   		
   		'KANAN
   		b21d3eaf-4e31-425c-ad1a-ba4e4002cacc Tool_Allocation_Numb_16,76
   		b21d3eaf-4e31-425c-ad1a-ba4e4002cacc Tool_Allocation_Numb_17,77
   		b21d3eaf-4e31-425c-ad1a-ba4e4002cacc Tool_Allocation_Numb_18,78
   		b21d3eaf-4e31-425c-ad1a-ba4e4002cacc Tool_Allocation_Numb_19,79
   		b21d3eaf-4e31-425c-ad1a-ba4e4002cacc Tool_Allocation_Numb_20,80
   		b21d3eaf-4e31-425c-ad1a-ba4e4002cacc Tool_Allocation_Numb_21,81
   		b21d3eaf-4e31-425c-ad1a-ba4e4002cacc Tool_Allocation_Numb_22,82
   		b21d3eaf-4e31-425c-ad1a-ba4e4002cacc Tool_Allocation_Numb_23,83
   		b21d3eaf-4e31-425c-ad1a-ba4e4002cacc Tool_Allocation_Numb_24,84
   		b21d3eaf-4e31-425c-ad1a-ba4e4002cacc Tool_Allocation_Numb_25,85
   		b21d3eaf-4e31-425c-ad1a-ba4e4002cacc Tool_Allocation_Numb_26,86
   		b21d3eaf-4e31-425c-ad1a-ba4e4002cacc Tool_Allocation_Numb_27,87
   		b21d3eaf-4e31-425c-ad1a-ba4e4002cacc Tool_Allocation_Numb_28,88
   		b21d3eaf-4e31-425c-ad1a-ba4e4002cacc Tool_Allocation_Numb_29,89
   		b21d3eaf-4e31-425c-ad1a-ba4e4002cacc Tool_Allocation_Numb_30,90		
   Case 4
   		b21d3eaf-4e31-425c-ad1a-ba4e4002cacc Tool_Allocation_Numb_1,91
   		b21d3eaf-4e31-425c-ad1a-ba4e4002cacc Tool_Allocation_Numb_2,92
   		b21d3eaf-4e31-425c-ad1a-ba4e4002cacc Tool_Allocation_Numb_3,93
   		b21d3eaf-4e31-425c-ad1a-ba4e4002cacc Tool_Allocation_Numb_4,94
   		b21d3eaf-4e31-425c-ad1a-ba4e4002cacc Tool_Allocation_Numb_5,95
   		b21d3eaf-4e31-425c-ad1a-ba4e4002cacc Tool_Allocation_Numb_6,96
   		b21d3eaf-4e31-425c-ad1a-ba4e4002cacc Tool_Allocation_Numb_7,97
   		b21d3eaf-4e31-425c-ad1a-ba4e4002cacc Tool_Allocation_Numb_8,98
   		b21d3eaf-4e31-425c-ad1a-ba4e4002cacc Tool_Allocation_Numb_9,99
   		b21d3eaf-4e31-425c-ad1a-ba4e4002cacc Tool_Allocation_Numb_10,100
   		b21d3eaf-4e31-425c-ad1a-ba4e4002cacc Tool_Allocation_Numb_11,101
   		b21d3eaf-4e31-425c-ad1a-ba4e4002cacc Tool_Allocation_Numb_12,102
   		b21d3eaf-4e31-425c-ad1a-ba4e4002cacc Tool_Allocation_Numb_13,103
   		b21d3eaf-4e31-425c-ad1a-ba4e4002cacc Tool_Allocation_Numb_14,104
   		b21d3eaf-4e31-425c-ad1a-ba4e4002cacc Tool_Allocation_Numb_15,105
   		
   		'KANAN
   		b21d3eaf-4e31-425c-ad1a-ba4e4002cacc Tool_Allocation_Numb_16,106
   		b21d3eaf-4e31-425c-ad1a-ba4e4002cacc Tool_Allocation_Numb_17,107
   		b21d3eaf-4e31-425c-ad1a-ba4e4002cacc Tool_Allocation_Numb_18,108
   		b21d3eaf-4e31-425c-ad1a-ba4e4002cacc Tool_Allocation_Numb_19,109
   		b21d3eaf-4e31-425c-ad1a-ba4e4002cacc Tool_Allocation_Numb_20,110
   		b21d3eaf-4e31-425c-ad1a-ba4e4002cacc Tool_Allocation_Numb_21,111
   		b21d3eaf-4e31-425c-ad1a-ba4e4002cacc Tool_Allocation_Numb_22,112
   		b21d3eaf-4e31-425c-ad1a-ba4e4002cacc Tool_Allocation_Numb_23,113
   		b21d3eaf-4e31-425c-ad1a-ba4e4002cacc Tool_Allocation_Numb_24,114
   		b21d3eaf-4e31-425c-ad1a-ba4e4002cacc Tool_Allocation_Numb_25,115
   		b21d3eaf-4e31-425c-ad1a-ba4e4002cacc Tool_Allocation_Numb_26,116
   		b21d3eaf-4e31-425c-ad1a-ba4e4002cacc Tool_Allocation_Numb_27,117
   		b21d3eaf-4e31-425c-ad1a-ba4e4002cacc Tool_Allocation_Numb_28,118
   		b21d3eaf-4e31-425c-ad1a-ba4e4002cacc Tool_Allocation_Numb_29,119
   		b21d3eaf-4e31-425c-ad1a-ba4e4002cacc Tool_Allocation_Numb_30,120		
   Case Else
   	'KIRI
   		
   		b21d3eaf-4e31-425c-ad1a-ba4e4002cacc Tool_Allocation_Numb_1,1
   		b21d3eaf-4e31-425c-ad1a-ba4e4002cacc Tool_Allocation_Numb_2,2
   		b21d3eaf-4e31-425c-ad1a-ba4e4002cacc Tool_Allocation_Numb_3,3
   		b21d3eaf-4e31-425c-ad1a-ba4e4002cacc Tool_Allocation_Numb_4,4
   		b21d3eaf-4e31-425c-ad1a-ba4e4002cacc Tool_Allocation_Numb_5,5
   		b21d3eaf-4e31-425c-ad1a-ba4e4002cacc Tool_Allocation_Numb_6,6
   		b21d3eaf-4e31-425c-ad1a-ba4e4002cacc Tool_Allocation_Numb_7,7
   		b21d3eaf-4e31-425c-ad1a-ba4e4002cacc Tool_Allocation_Numb_8,8
   		b21d3eaf-4e31-425c-ad1a-ba4e4002cacc Tool_Allocation_Numb_9,9
   		b21d3eaf-4e31-425c-ad1a-ba4e4002cacc Tool_Allocation_Numb_10,10
   		b21d3eaf-4e31-425c-ad1a-ba4e4002cacc Tool_Allocation_Numb_11,11
   		b21d3eaf-4e31-425c-ad1a-ba4e4002cacc Tool_Allocation_Numb_12,12
   		b21d3eaf-4e31-425c-ad1a-ba4e4002cacc Tool_Allocation_Numb_13,13
   		b21d3eaf-4e31-425c-ad1a-ba4e4002cacc Tool_Allocation_Numb_14,14
   		b21d3eaf-4e31-425c-ad1a-ba4e4002cacc Tool_Allocation_Numb_15,15
   		
   		'KANAN
   		b21d3eaf-4e31-425c-ad1a-ba4e4002cacc Tool_Allocation_Numb_16,16
   		b21d3eaf-4e31-425c-ad1a-ba4e4002cacc Tool_Allocation_Numb_17,17
   		b21d3eaf-4e31-425c-ad1a-ba4e4002cacc Tool_Allocation_Numb_18,18
   		b21d3eaf-4e31-425c-ad1a-ba4e4002cacc Tool_Allocation_Numb_19,19
   		b21d3eaf-4e31-425c-ad1a-ba4e4002cacc Tool_Allocation_Numb_20,20
   		b21d3eaf-4e31-425c-ad1a-ba4e4002cacc Tool_Allocation_Numb_21,21
   		b21d3eaf-4e31-425c-ad1a-ba4e4002cacc Tool_Allocation_Numb_22,22
   		b21d3eaf-4e31-425c-ad1a-ba4e4002cacc Tool_Allocation_Numb_23,23
   		b21d3eaf-4e31-425c-ad1a-ba4e4002cacc Tool_Allocation_Numb_24,24
   		b21d3eaf-4e31-425c-ad1a-ba4e4002cacc Tool_Allocation_Numb_25,25
   		b21d3eaf-4e31-425c-ad1a-ba4e4002cacc Tool_Allocation_Numb_26,26
   		b21d3eaf-4e31-425c-ad1a-ba4e4002cacc Tool_Allocation_Numb_27,27
   		b21d3eaf-4e31-425c-ad1a-ba4e4002cacc Tool_Allocation_Numb_28,28
   		b21d3eaf-4e31-425c-ad1a-ba4e4002cacc Tool_Allocation_Numb_29,29
   		b21d3eaf-4e31-425c-ad1a-ba4e4002cacc Tool_Allocation_Numb_30,30			
   End Select
   		

VB script "ToolAllocation_Sec"
   'Tip:
   ' 1. Use the <CTRL+SPACE> or <CTRL+I> shortcut to open a list of all objects and functions
   ' 2. Write the code using the HMI Runtime object.
   '  Example: HmiRuntime.Screens("Screen_1").
   ' 3. Use the <CTRL+J> shortcut to create an object reference.
   'Write the code as of this position:
    If SmartTags("DB939_Tool_alloc_HMI_Limit_allocation_list")<30 Then
   	 b21d3eaf-4e31-425c-ad1a-ba4e4002cacc Tool_Allocation_Numb_1,1
   		b21d3eaf-4e31-425c-ad1a-ba4e4002cacc Tool_Allocation_Numb_2,2
   		b21d3eaf-4e31-425c-ad1a-ba4e4002cacc Tool_Allocation_Numb_3,3
   		b21d3eaf-4e31-425c-ad1a-ba4e4002cacc Tool_Allocation_Numb_4,4
   		b21d3eaf-4e31-425c-ad1a-ba4e4002cacc Tool_Allocation_Numb_5,5
   		b21d3eaf-4e31-425c-ad1a-ba4e4002cacc Tool_Allocation_Numb_6,6
   		b21d3eaf-4e31-425c-ad1a-ba4e4002cacc Tool_Allocation_Numb_7,7
   		b21d3eaf-4e31-425c-ad1a-ba4e4002cacc Tool_Allocation_Numb_8,8
   		b21d3eaf-4e31-425c-ad1a-ba4e4002cacc Tool_Allocation_Numb_9,9
   		b21d3eaf-4e31-425c-ad1a-ba4e4002cacc Tool_Allocation_Numb_10,10
   		b21d3eaf-4e31-425c-ad1a-ba4e4002cacc Tool_Allocation_Numb_11,11
   		b21d3eaf-4e31-425c-ad1a-ba4e4002cacc Tool_Allocation_Numb_12,12
   		b21d3eaf-4e31-425c-ad1a-ba4e4002cacc Tool_Allocation_Numb_13,13
   		b21d3eaf-4e31-425c-ad1a-ba4e4002cacc Tool_Allocation_Numb_14,14
   		b21d3eaf-4e31-425c-ad1a-ba4e4002cacc Tool_Allocation_Numb_15,15
   		
   		'KANAN
   		b21d3eaf-4e31-425c-ad1a-ba4e4002cacc Tool_Allocation_Numb_16,16
   		b21d3eaf-4e31-425c-ad1a-ba4e4002cacc Tool_Allocation_Numb_17,17
   		b21d3eaf-4e31-425c-ad1a-ba4e4002cacc Tool_Allocation_Numb_18,18
   		b21d3eaf-4e31-425c-ad1a-ba4e4002cacc Tool_Allocation_Numb_19,19
   		b21d3eaf-4e31-425c-ad1a-ba4e4002cacc Tool_Allocation_Numb_20,20
   		b21d3eaf-4e31-425c-ad1a-ba4e4002cacc Tool_Allocation_Numb_21,21
   		b21d3eaf-4e31-425c-ad1a-ba4e4002cacc Tool_Allocation_Numb_22,22
   		b21d3eaf-4e31-425c-ad1a-ba4e4002cacc Tool_Allocation_Numb_23,23
   		b21d3eaf-4e31-425c-ad1a-ba4e4002cacc Tool_Allocation_Numb_24,24
   		b21d3eaf-4e31-425c-ad1a-ba4e4002cacc Tool_Allocation_Numb_25,25
   		b21d3eaf-4e31-425c-ad1a-ba4e4002cacc Tool_Allocation_Numb_26,26
   		b21d3eaf-4e31-425c-ad1a-ba4e4002cacc Tool_Allocation_Numb_27,27
   		b21d3eaf-4e31-425c-ad1a-ba4e4002cacc Tool_Allocation_Numb_28,28
   		b21d3eaf-4e31-425c-ad1a-ba4e4002cacc Tool_Allocation_Numb_29,29
   		b21d3eaf-4e31-425c-ad1a-ba4e4002cacc Tool_Allocation_Numb_30,30		
   
   End If
    

VB script "Consumtion"
   Select Case SmartTags("DB_Zaehler_Anzeige_ReadWriteDeviceNo")
   	
   	Case 1:
   		b21d3eaf-4e31-425c-ad1a-ba4e4002cacc Consumtion_Numb_1,1
   		b21d3eaf-4e31-425c-ad1a-ba4e4002cacc Consumtion_Numb_2,2
   		b21d3eaf-4e31-425c-ad1a-ba4e4002cacc Consumtion_Numb_3,3
   		b21d3eaf-4e31-425c-ad1a-ba4e4002cacc Consumtion_Numb_4,4
   		b21d3eaf-4e31-425c-ad1a-ba4e4002cacc Consumtion_Numb_5,5
   		b21d3eaf-4e31-425c-ad1a-ba4e4002cacc Consumtion_Numb_6,6
   		b21d3eaf-4e31-425c-ad1a-ba4e4002cacc Consumtion_Numb_7,7
   		b21d3eaf-4e31-425c-ad1a-ba4e4002cacc Consumtion_Numb_8,8
   		b21d3eaf-4e31-425c-ad1a-ba4e4002cacc Consumtion_Numb_9,9
   		b21d3eaf-4e31-425c-ad1a-ba4e4002cacc Consumtion_Numb_10,10
   	Case 11:
   		b21d3eaf-4e31-425c-ad1a-ba4e4002cacc Consumtion_Numb_1,11
   		b21d3eaf-4e31-425c-ad1a-ba4e4002cacc Consumtion_Numb_2,12
   		b21d3eaf-4e31-425c-ad1a-ba4e4002cacc Consumtion_Numb_3,13
   		b21d3eaf-4e31-425c-ad1a-ba4e4002cacc Consumtion_Numb_4,14
   		b21d3eaf-4e31-425c-ad1a-ba4e4002cacc Consumtion_Numb_5,15
   		b21d3eaf-4e31-425c-ad1a-ba4e4002cacc Consumtion_Numb_6,16
   		b21d3eaf-4e31-425c-ad1a-ba4e4002cacc Consumtion_Numb_7,17
   		b21d3eaf-4e31-425c-ad1a-ba4e4002cacc Consumtion_Numb_8,18
   		b21d3eaf-4e31-425c-ad1a-ba4e4002cacc Consumtion_Numb_9,19
   		b21d3eaf-4e31-425c-ad1a-ba4e4002cacc Consumtion_Numb_10,20	
   	Case 21:
   		b21d3eaf-4e31-425c-ad1a-ba4e4002cacc Consumtion_Numb_1,21
   		b21d3eaf-4e31-425c-ad1a-ba4e4002cacc Consumtion_Numb_2,22
   		b21d3eaf-4e31-425c-ad1a-ba4e4002cacc Consumtion_Numb_3,23
   		b21d3eaf-4e31-425c-ad1a-ba4e4002cacc Consumtion_Numb_4,24
   		b21d3eaf-4e31-425c-ad1a-ba4e4002cacc Consumtion_Numb_5,25
   		b21d3eaf-4e31-425c-ad1a-ba4e4002cacc Consumtion_Numb_6,26
   		b21d3eaf-4e31-425c-ad1a-ba4e4002cacc Consumtion_Numb_7,27
   		b21d3eaf-4e31-425c-ad1a-ba4e4002cacc Consumtion_Numb_8,28
   		b21d3eaf-4e31-425c-ad1a-ba4e4002cacc Consumtion_Numb_9,29
   		b21d3eaf-4e31-425c-ad1a-ba4e4002cacc Consumtion_Numb_10,30
   	
   	Case 31:
   		b21d3eaf-4e31-425c-ad1a-ba4e4002cacc Consumtion_Numb_1,31
   		b21d3eaf-4e31-425c-ad1a-ba4e4002cacc Consumtion_Numb_2,32
   		b21d3eaf-4e31-425c-ad1a-ba4e4002cacc Consumtion_Numb_3,33
   		b21d3eaf-4e31-425c-ad1a-ba4e4002cacc Consumtion_Numb_4,34
   		b21d3eaf-4e31-425c-ad1a-ba4e4002cacc Consumtion_Numb_5,35
   		b21d3eaf-4e31-425c-ad1a-ba4e4002cacc Consumtion_Numb_6,36
   		b21d3eaf-4e31-425c-ad1a-ba4e4002cacc Consumtion_Numb_7,37
   		b21d3eaf-4e31-425c-ad1a-ba4e4002cacc Consumtion_Numb_8,38
   		b21d3eaf-4e31-425c-ad1a-ba4e4002cacc Consumtion_Numb_9,39
   		b21d3eaf-4e31-425c-ad1a-ba4e4002cacc Consumtion_Numb_10,40
   	Case 41:
   		b21d3eaf-4e31-425c-ad1a-ba4e4002cacc Consumtion_Numb_1,41
   		b21d3eaf-4e31-425c-ad1a-ba4e4002cacc Consumtion_Numb_2,42
   		b21d3eaf-4e31-425c-ad1a-ba4e4002cacc Consumtion_Numb_3,43
   		b21d3eaf-4e31-425c-ad1a-ba4e4002cacc Consumtion_Numb_4,44
   		b21d3eaf-4e31-425c-ad1a-ba4e4002cacc Consumtion_Numb_5,45
   		b21d3eaf-4e31-425c-ad1a-ba4e4002cacc Consumtion_Numb_6,46
   		b21d3eaf-4e31-425c-ad1a-ba4e4002cacc Consumtion_Numb_7,47
   		b21d3eaf-4e31-425c-ad1a-ba4e4002cacc Consumtion_Numb_8,48
   		b21d3eaf-4e31-425c-ad1a-ba4e4002cacc Consumtion_Numb_9,49
   		b21d3eaf-4e31-425c-ad1a-ba4e4002cacc Consumtion_Numb_10,50
   	Case 51:
   		b21d3eaf-4e31-425c-ad1a-ba4e4002cacc Consumtion_Numb_1,51
   		b21d3eaf-4e31-425c-ad1a-ba4e4002cacc Consumtion_Numb_2,52
   		b21d3eaf-4e31-425c-ad1a-ba4e4002cacc Consumtion_Numb_3,53
   		b21d3eaf-4e31-425c-ad1a-ba4e4002cacc Consumtion_Numb_4,54
   		b21d3eaf-4e31-425c-ad1a-ba4e4002cacc Consumtion_Numb_5,55
   		b21d3eaf-4e31-425c-ad1a-ba4e4002cacc Consumtion_Numb_6,56
   		b21d3eaf-4e31-425c-ad1a-ba4e4002cacc Consumtion_Numb_7,57
   		b21d3eaf-4e31-425c-ad1a-ba4e4002cacc Consumtion_Numb_8,58
   		b21d3eaf-4e31-425c-ad1a-ba4e4002cacc Consumtion_Numb_9,59
   		b21d3eaf-4e31-425c-ad1a-ba4e4002cacc Consumtion_Numb_10,60
   	Case Else:
   		b21d3eaf-4e31-425c-ad1a-ba4e4002cacc Consumtion_Numb_1,1
   		b21d3eaf-4e31-425c-ad1a-ba4e4002cacc Consumtion_Numb_2,2
   		b21d3eaf-4e31-425c-ad1a-ba4e4002cacc Consumtion_Numb_3,3
   		b21d3eaf-4e31-425c-ad1a-ba4e4002cacc Consumtion_Numb_4,4
   		b21d3eaf-4e31-425c-ad1a-ba4e4002cacc Consumtion_Numb_5,5
   		b21d3eaf-4e31-425c-ad1a-ba4e4002cacc Consumtion_Numb_6,6
   		b21d3eaf-4e31-425c-ad1a-ba4e4002cacc Consumtion_Numb_7,7
   		b21d3eaf-4e31-425c-ad1a-ba4e4002cacc Consumtion_Numb_8,8
   		b21d3eaf-4e31-425c-ad1a-ba4e4002cacc Consumtion_Numb_9,9
   		b21d3eaf-4e31-425c-ad1a-ba4e4002cacc Consumtion_Numb_10,10
   End Select

VB script "Consumtion_Increase"
   If SmartTags("DB_Zaehler_Anzeige_ReadWriteDeviceNo") < 51 Then
   	SmartTags("DB_Zaehler_Anzeige_ReadWriteDeviceNo")=SmartTags("DB_Zaehler_Anzeige_ReadWriteDeviceNo")+10
   End If

VB script "Consumtiom_Decrease"
    If SmartTags("DB_Zaehler_Anzeige_ReadWriteDeviceNo") > 1 Then
   	 SmartTags("DB_Zaehler_Anzeige_ReadWriteDeviceNo")=SmartTags("DB_Zaehler_Anzeige_ReadWriteDeviceNo")-10
    end if
    

VB script "PopUp_ToolEditor"
   If SmartTags("DB_MouldEditor_HMI_uData_sStatusBits_xFaultDeleteProgram")=True Then
   	efd93a16-2665-4b85-bcb9-25eddcb7b6f4 Save,446,387,$3$hmiToggle$,$3$hmiAnimationOff$,$3$hmiSlow$
   		
   End If

VB script "VBStore_tool"
   Dim fs, f, FName, Header, ToolNo, ToolName, PSno, PS, RefComp, MH, ShotTime, TotalFlow,	TotalWeight, PartCounter, Service, CP, Purge
   Dim Comp1, Comp2, Comp3, Comp4, Comp5, Comp6, FR1, FR2, FR3, FR4, FR5, FR6, Press1, Press2, Press3, Press4, Press5, Press6
   Dim Del
   
   ToolNo = SmartTags("DB_MouldEditor_HMI_uData_sSelected_iTool")
   ToolName = SmartTags("DB_MouldEditor_HMI_uData_uTools_tool_name")
   PSno = SmartTags("DB_MouldEditor_HMI_uData_uTools_PartShot_Amount")
   Del = SmartTags("DB930_Tools_Tool{"& ToolNo &"}_tool_name")
   
   On Error Resume Next
    ' FileSystemObject erstellen
    ' Create FileSystemObject
   Set fs = CreateObject("FileCtl.FileSystem") 
   
   ' FileObject erstellen
   ' Create FileObject
    Set f = CreateObject("FileCtl.File")
   fs.kill StoragePath & "\Tools\" & CStr(ToolNo) & "_*.csv"
   bfde4b54-0db7-4817-8032-87127bf19bb9 "VBStore_tool: Tool deleted: " & CStr(ToolNo) & "_*.csv"
   
   For PS = 1 To 8
   RefComp = SmartTags("DB_MouldEditor_HMI_uData_arShotSet{"& PS &"}_RefComponent")
   MH = SmartTags("DB_MouldEditor_HMI_uData_arShotSet{"& PS &"}_MHNo")
   ShotTime = SmartTags("DB_MouldEditor_HMI_uData_arShotSet{"& PS &"}_FoamingTime")
   TotalFlow = SmartTags("DB_MouldEditor_HMI_uData_sCalculatedValues_arTotalFlow{"& PS &"}")
   TotalWeight = SmartTags("DB_MouldEditor_HMI_uData_arShotSet{"& PS &"}_PartWeight")
   PartCounter = SmartTags("DB_MouldEditor_HMI_uData_arShotSet{"& PS &"}_PartCounter")
   Service = SmartTags("DB_MouldEditor_HMI_uData_arShotSet{"& PS &"}_PartShotDisable")
   CP = SmartTags("DB_MouldEditor_HMI_uData_arShotSet{"& PS &"}_CPMoveAfterShot")
   Purge = SmartTags("DB_MouldEditor_HMI_uData_arShotSet{"& PS &"}_PurgeMHAfterShot")
   Comp1 = SmartTags("DB753_MeteringPump_Pump{1}_Name")
   Comp2 = SmartTags("DB753_MeteringPump_Pump{2}_Name")
   Comp3 = SmartTags("DB753_MeteringPump_Pump{3}_Name")
   Comp4 = SmartTags("DB753_MeteringPump_Pump{4}_Name")
   Comp5 = SmartTags("DB753_MeteringPump_Pump{5}_Name")
   Comp6 = SmartTags("DB753_MeteringPump_Pump{6}_Name")
   FR1 = SmartTags("DB_MouldEditor_HMI_uData_arShotSet{"& PS &"}_Flow{1}")
   FR2 = SmartTags("DB_MouldEditor_HMI_uData_arShotSet{"& PS &"}_Flow{2}")
   FR3 = SmartTags("DB_MouldEditor_HMI_uData_arShotSet{"& PS &"}_Flow{3}")
   FR4 = SmartTags("DB_MouldEditor_HMI_uData_arShotSet{"& PS &"}_Flow{4}")
   FR5 = SmartTags("DB_MouldEditor_HMI_uData_arShotSet{"& PS &"}_Flow{5}")
   FR6 = SmartTags("DB_MouldEditor_HMI_uData_arShotSet{"& PS &"}_Flow{6}")
   Press1 = SmartTags("DB_MouldEditor_HMI_uData_arShotSet{"& PS &"}_Pressure{1}")
   Press2 = SmartTags("DB_MouldEditor_HMI_uData_arShotSet{"& PS &"}_Pressure{2}")
   Press3 = SmartTags("DB_MouldEditor_HMI_uData_arShotSet{"& PS &"}_Pressure{3}")
   Press4 = SmartTags("DB_MouldEditor_HMI_uData_arShotSet{"& PS &"}_Pressure{4}")
   Press5 = SmartTags("DB_MouldEditor_HMI_uData_arShotSet{"& PS &"}_Pressure{5}")
   Press6 = SmartTags("DB_MouldEditor_HMI_uData_arShotSet{"& PS &"}_Pressure{6}")
   ' Archivierungspfad (Eingangsparameter) und Dateiname zusammensetzen 
   ' Combine archivepath (input parameter) and filename
   FName = StoragePath & "\Tools\" & CStr(ToolNo) & "_" & CStr(ToolName) & ".csv" 
   
   ' Tabellenkopf zusammenstellen 
   ' Create table header 
    Header = "Part shot;RefComp;MH;Shot time;total flow;total weight;Part counter;Service;CP;Purge after shot"
   
   ' Datei öffnen bzw. erstellen, wenn sie noch nicht existiert.
   ' Open File or create file if it does not exist 
    f.open FName, 8 								
   
   ' Wenn Datei 0 Byte groß, dann ist sie neu
   ' If file is 0 byte the file is new
    If fs.FileLen(FName) = 0 Then 
   	 f.lineprint("Tool No.:;" & CStr(ToolNo))' & Chr(10))
   	 f.lineprint("Tool Name:;" & CStr(ToolName))' & Chr(10))
   	 f.lineprint("Part shots:;" & CStr(PSno))' & Chr(10))
   	 f.lineprint(Header)' & Chr(10)
   ' =0 => Tabellenkopf muss eingefügt werden
   ' =0 => Table header must be inserted
    End If
   
   ' Werte der Variablen in die Archivdatei schreiben (Parameter "TagName" z.B. Tag_01)
   ' Write values of variables in archive file (Parameter "TagName" for sample Tag_01)
    f.lineprint(CStr(PS) & ";" & CStr(RefComp) & ";" & CStr(MH) & ";" & CStr(ShotTime) & ";" & CStr(TotalFlow) & ";" & CStr(TotalWeight) & ";" & CStr(PartCounter) & ";" & CStr(Service) & ";" & CStr(CP) & ";" & CStr(Purge))' & Chr(10)
    f.lineprint("Component name:;" & CStr(Comp1) & ";" & CStr(Comp2) & ";" & CStr(Comp3) & ";" & CStr(Comp4) & ";" & CStr(Comp5) & ";" & CStr(Comp6))' & Chr(10))
    f.lineprint("Flow rate:;" & CStr(FR1) & ";" & CStr(FR2) & ";" & CStr(FR3) & ";" & CStr(FR4) & ";" & CStr(FR5) & ";" & CStr(FR6))' & Chr(10))
    f.lineprint("Pressure::;" & CStr(Press1) & ";" & CStr(Press2) & ";" & CStr(Press3) & ";" & CStr(Press4) & ";" & CStr(Press5) & ";" & CStr(Press6))' & Chr(10))
    f.lineprint("--------------------")
   ' Datei wieder schließen
   ' Close file
    f.Close
   
   
   Next
   
   ' Verwendeten Speicher wieder freigeben
   ' Used storage will be freed
   Set f  = Nothing
   Set fs = Nothing
   'ShowSystemAlarm "comp " & PS
   
   'Error checking
   If Err.Number <>0 Then
   bfde4b54-0db7-4817-8032-87127bf19bb9 "Error#" & CStr(Err.Number) & " " & Err.Description
   Err.Clear
   ' Exit Sub'
   End If
   
   bfde4b54-0db7-4817-8032-87127bf19bb9 "VBStore_tool: " & CStr(ToolNo) & "_" & CStr(ToolName) & ".csv"

VB script "VBStore_tool_Deleted"
   Dim fs, f, FName, Header, ToolNo, ToolName, PSno
   Dim Del
   
   ToolNo = SmartTags("DB_MouldEditor_HMI_uData_sSelected_iTool")
   ToolName = SmartTags("DB_MouldEditor_HMI_uData_uTools_tool_name")
   PSno = SmartTags("DB_MouldEditor_HMI_uData_uTools_PartShot_Amount")
   Del = SmartTags("DB930_Tools_Tool{"& ToolNo &"}_tool_name")
   
   
   f38ba6b2-0c13-4a6f-acab-73f2fde9baea 1,SmartTags("DB_MouldEditor_HMI_uData_sSelected_iTool"),$3$hmiOverwriteAlways$,$3$hmiOff$,Null 
   
   
   On Error Resume Next
    ' FileSystemObject erstellen
    ' Create FileSystemObject
   Set fs = CreateObject("FileCtl.FileSystem") 
   
   ' FileObject erstellen
   ' Create FileObject
    Set f = CreateObject("FileCtl.File")
   fs.kill StoragePath & "\Tools\" & CStr(ToolNo) & "_"& CStr(ToolName) & ".csv"
   bfde4b54-0db7-4817-8032-87127bf19bb9 "VBStore_tool: Tool deleted: " & CStr(ToolNo) & "_" & CStr(ToolName) & ".csv"
   
   ' Verwendeten Speicher wieder freigeben
   ' Used storage will be freed
   Set f  = Nothing
   Set fs = Nothing
   'ShowSystemAlarm "comp " & PS
   
   
   'Error checking
   If Err.Number <>0 Then
   bfde4b54-0db7-4817-8032-87127bf19bb9 "Error#" & CStr(Err.Number) & " " & Err.Description
   Err.Clear
   ' Exit Sub'
   End If
   
   bfde4b54-0db7-4817-8032-87127bf19bb9 "Data record no. " & CStr(ToolNo) & " has been successfully saved."

VB script "ReadDataFromSD"
   '/////////////////////////////////////////////////////////////////////////
   ' en: Script for the readout of a text file      
   ' de: Skript zum Auslesen einer Textdatei
   ' Created: 29-05-2007
   ' Version: v0.1
   ' Author:  ZW										   only for Windows CE
   '/////////////////////////////////////////////////////////////////////////
   
   'Declaration of local tags - Deklaration von lokalen Variablen
   Dim f, path, MyZf, i, j, field, HiField(43,10), PS, Je, Flo, Pre
   
   'If bExtension = 0 Then
   	'path = "\flash\textfile.txt"
   '	path = "\Storage Card2\textfile.txt"
   'Else
   	'path = "\flash\textfile.csv"
   	path = SmartTags("ImportDataFrom_SD") '"\Storage Card2\textfile.csv"
   'End If
   
   'Error Routine - Fehlerroutine
   On Error Resume Next
   
   If SmartTags("ImportDataFrom_SD_stat")= 0 Then
   	'Create object - Objekt erstellen
   Set f = CreateObject("FileCtl.File")
   
   If Err.Number <> 0 Then
   	bfde4b54-0db7-4817-8032-87127bf19bb9 "Error #" & CStr(Err.Number) & " " & Err.Description
   	Err.Clear
   	Exit Sub
   End If
   
   'Open file - Datei öffnen
   f.open path, 1
   
   If Err.Number <> 0 Then
   	bfde4b54-0db7-4817-8032-87127bf19bb9 "Error #" & CStr(Err.Number) & " " & Err.Description
   	Err.Clear
   	Exit Sub
   End If
   
   'Loop
   Do While f.EOF = False
   	MyZf = f.LineInputString
   	field = Split(MyZf, ";")
   	
   	For i=0 To 43
   		field(i) = Replace(field(i), " ", "")
   		HiField(j,i) = field(i)
   	Next
   	
   	SmartTags("DB_MouldEditor_HMI_uData_uTools_tool_name") = HiField(1,1)
   	SmartTags("DB_MouldEditor_HMI_uData_uTools_PartShot_Amount") = HiField(2,1)
   	
   	SmartTags("DB_MouldEditor_HMI_uData_arShotSet{1}_RefComponent") = HiField(4,1)
   	SmartTags("DB_MouldEditor_HMI_uData_arShotSet{1}_MHNo") = HiField(4,2)
   	SmartTags("DB_MouldEditor_HMI_uData_arShotSet{1}_FoamingTime") = HiField(4,3)
   	SmartTags("DB_MouldEditor_HMI_uData_sCalculatedValues_arTotalFlow{1}") = HiField(4,4)
   	SmartTags("DB_MouldEditor_HMI_uData_arShotSet{1}_PartWeight") = HiField(4,5)
   	SmartTags("DB_MouldEditor_HMI_uData_arShotSet{1}_PartCounter") = HiField(4,6)
   	SmartTags("DB_MouldEditor_HMI_uData_arShotSet{1}_PartShotDisable") = HiField(4,7)
   	SmartTags("DB_MouldEditor_HMI_uData_arShotSet{1}_CPMoveAfterShot") = HiField(4,8)
   	SmartTags("DB_MouldEditor_HMI_uData_arShotSet{1}_PurgeMHAfterShot") = HiField(4,9)
   	
   	SmartTags("DB_MouldEditor_HMI_uData_arShotSet{2}_RefComponent") = HiField(9,1)
   	SmartTags("DB_MouldEditor_HMI_uData_arShotSet{2}_MHNo") = HiField(9,2)
   	SmartTags("DB_MouldEditor_HMI_uData_arShotSet{2}_FoamingTime") = HiField(9,3)
   	SmartTags("DB_MouldEditor_HMI_uData_sCalculatedValues_arTotalFlow{2}") = HiField(9,4)
   	SmartTags("DB_MouldEditor_HMI_uData_arShotSet{2}_PartWeight") = HiField(9,5)
   	SmartTags("DB_MouldEditor_HMI_uData_arShotSet{2}_PartCounter") = HiField(9,6)
   	SmartTags("DB_MouldEditor_HMI_uData_arShotSet{2}_PartShotDisable") = HiField(9,7)
   	SmartTags("DB_MouldEditor_HMI_uData_arShotSet{2}_CPMoveAfterShot") = HiField(9,8)
   	SmartTags("DB_MouldEditor_HMI_uData_arShotSet{2}_PurgeMHAfterShot") = HiField(9,9)
   	
   	SmartTags("DB_MouldEditor_HMI_uData_arShotSet{3}_RefComponent") = HiField(14,1)
   	SmartTags("DB_MouldEditor_HMI_uData_arShotSet{3}_MHNo") = HiField(14,2)
   	SmartTags("DB_MouldEditor_HMI_uData_arShotSet{3}_FoamingTime") = HiField(14,3)
   	SmartTags("DB_MouldEditor_HMI_uData_sCalculatedValues_arTotalFlow{3}") = HiField(14,4)
   	SmartTags("DB_MouldEditor_HMI_uData_arShotSet{3}_PartWeight") = HiField(14,5)
   	SmartTags("DB_MouldEditor_HMI_uData_arShotSet{3}_PartCounter") = HiField(14,6)
   	SmartTags("DB_MouldEditor_HMI_uData_arShotSet{3}_PartShotDisable") = HiField(14,7)
   	SmartTags("DB_MouldEditor_HMI_uData_arShotSet{3}_CPMoveAfterShot") = HiField(14,8)
   	SmartTags("DB_MouldEditor_HMI_uData_arShotSet{3}_PurgeMHAfterShot") = HiField(14,9)
   	
   	SmartTags("DB_MouldEditor_HMI_uData_arShotSet{4}_RefComponent") = HiField(19,1)
   	SmartTags("DB_MouldEditor_HMI_uData_arShotSet{4}_MHNo") = HiField(19,2)
   	SmartTags("DB_MouldEditor_HMI_uData_arShotSet{4}_FoamingTime") = HiField(19,3)
   	SmartTags("DB_MouldEditor_HMI_uData_sCalculatedValues_arTotalFlow{4}") = HiField(19,4)
   	SmartTags("DB_MouldEditor_HMI_uData_arShotSet{4}_PartWeight") = HiField(19,5)
   	SmartTags("DB_MouldEditor_HMI_uData_arShotSet{4}_PartCounter") = HiField(19,6)
   	SmartTags("DB_MouldEditor_HMI_uData_arShotSet{4}_PartShotDisable") = HiField(19,7)
   	SmartTags("DB_MouldEditor_HMI_uData_arShotSet{4}_CPMoveAfterShot") = HiField(19,8)
   	SmartTags("DB_MouldEditor_HMI_uData_arShotSet{4}_PurgeMHAfterShot") = HiField(19,9)
   	
   	SmartTags("DB_MouldEditor_HMI_uData_arShotSet{5}_RefComponent") = HiField(24,1)
   	SmartTags("DB_MouldEditor_HMI_uData_arShotSet{5}_MHNo") = HiField(24,2)
   	SmartTags("DB_MouldEditor_HMI_uData_arShotSet{5}_FoamingTime") = HiField(24,3)
   	SmartTags("DB_MouldEditor_HMI_uData_sCalculatedValues_arTotalFlow{5}") = HiField(24,4)
   	SmartTags("DB_MouldEditor_HMI_uData_arShotSet{5}_PartWeight") = HiField(24,5)
   	SmartTags("DB_MouldEditor_HMI_uData_arShotSet{5}_PartCounter") = HiField(24,6)
   	SmartTags("DB_MouldEditor_HMI_uData_arShotSet{5}_PartShotDisable") = HiField(24,7)
   	SmartTags("DB_MouldEditor_HMI_uData_arShotSet{5}_CPMoveAfterShot") = HiField(24,8)
   	SmartTags("DB_MouldEditor_HMI_uData_arShotSet{5}_PurgeMHAfterShot") = HiField(24,9)
   	
   	SmartTags("DB_MouldEditor_HMI_uData_arShotSet{6}_RefComponent") = HiField(29,1)
   	SmartTags("DB_MouldEditor_HMI_uData_arShotSet{6}_MHNo") = HiField(29,2)
   	SmartTags("DB_MouldEditor_HMI_uData_arShotSet{6}_FoamingTime") = HiField(29,3)
   	SmartTags("DB_MouldEditor_HMI_uData_sCalculatedValues_arTotalFlow{6}") = HiField(29,4)
   	SmartTags("DB_MouldEditor_HMI_uData_arShotSet{6}_PartWeight") = HiField(29,5)
   	SmartTags("DB_MouldEditor_HMI_uData_arShotSet{6}_PartCounter") = HiField(29,6)
   	SmartTags("DB_MouldEditor_HMI_uData_arShotSet{6}_PartShotDisable") = HiField(29,7)
   	SmartTags("DB_MouldEditor_HMI_uData_arShotSet{6}_CPMoveAfterShot") = HiField(29,8)
   	SmartTags("DB_MouldEditor_HMI_uData_arShotSet{6}_PurgeMHAfterShot") = HiField(29,9)
   	
   	SmartTags("DB_MouldEditor_HMI_uData_arShotSet{7}_RefComponent") = HiField(34,1)
   	SmartTags("DB_MouldEditor_HMI_uData_arShotSet{7}_MHNo") = HiField(34,2)
   	SmartTags("DB_MouldEditor_HMI_uData_arShotSet{7}_FoamingTime") = HiField(34,3)
   	SmartTags("DB_MouldEditor_HMI_uData_sCalculatedValues_arTotalFlow{7}") = HiField(34,4)
   	SmartTags("DB_MouldEditor_HMI_uData_arShotSet{7}_PartWeight") = HiField(34,5)
   	SmartTags("DB_MouldEditor_HMI_uData_arShotSet{7}_PartCounter") = HiField(34,6)
   	SmartTags("DB_MouldEditor_HMI_uData_arShotSet{7}_PartShotDisable") = HiField(34,7)
   	SmartTags("DB_MouldEditor_HMI_uData_arShotSet{7}_CPMoveAfterShot") = HiField(34,8)
   	SmartTags("DB_MouldEditor_HMI_uData_arShotSet{7}_PurgeMHAfterShot") = HiField(34,9)
   	
   	SmartTags("DB_MouldEditor_HMI_uData_arShotSet{8}_RefComponent") = HiField(39,1)
   	SmartTags("DB_MouldEditor_HMI_uData_arShotSet{8}_MHNo") = HiField(39,2)
   	SmartTags("DB_MouldEditor_HMI_uData_arShotSet{8}_FoamingTime") = HiField(39,3)
   	SmartTags("DB_MouldEditor_HMI_uData_sCalculatedValues_arTotalFlow{8}") = HiField(39,4)
   	SmartTags("DB_MouldEditor_HMI_uData_arShotSet{8}_PartWeight") = HiField(39,5)
   	SmartTags("DB_MouldEditor_HMI_uData_arShotSet{8}_PartCounter") = HiField(39,6)
   	SmartTags("DB_MouldEditor_HMI_uData_arShotSet{8}_PartShotDisable") = HiField(39,7)
   	SmartTags("DB_MouldEditor_HMI_uData_arShotSet{8}_CPMoveAfterShot") = HiField(39,8)
   	SmartTags("DB_MouldEditor_HMI_uData_arShotSet{8}_PurgeMHAfterShot") = HiField(39,9)
   	
   	'//FLOW
   	SmartTags("DB_MouldEditor_HMI_uData_arShotSet{1}_Flow{1}")=HiField(6,1)
   	SmartTags("DB_MouldEditor_HMI_uData_arShotSet{1}_Flow{2}")=HiField(6,2)	
   	SmartTags("DB_MouldEditor_HMI_uData_arShotSet{1}_Flow{3}")=HiField(6,3)
   	SmartTags("DB_MouldEditor_HMI_uData_arShotSet{1}_Flow{4}")=HiField(6,4)
   	SmartTags("DB_MouldEditor_HMI_uData_arShotSet{1}_Flow{5}")=HiField(6,5)	
   	SmartTags("DB_MouldEditor_HMI_uData_arShotSet{1}_Flow{6}")=HiField(6,6)
   	
   	SmartTags("DB_MouldEditor_HMI_uData_arShotSet{2}_Flow{1}")=HiField(11,1)
   	SmartTags("DB_MouldEditor_HMI_uData_arShotSet{2}_Flow{2}")=HiField(11,2)	
   	SmartTags("DB_MouldEditor_HMI_uData_arShotSet{2}_Flow{3}")=HiField(11,3)
   	SmartTags("DB_MouldEditor_HMI_uData_arShotSet{2}_Flow{4}")=HiField(11,4)
   	SmartTags("DB_MouldEditor_HMI_uData_arShotSet{2}_Flow{5}")=HiField(11,5)	
   	SmartTags("DB_MouldEditor_HMI_uData_arShotSet{2}_Flow{6}")=HiField(11,6)
   	
   	SmartTags("DB_MouldEditor_HMI_uData_arShotSet{3}_Flow{1}")=HiField(16,1)
   	SmartTags("DB_MouldEditor_HMI_uData_arShotSet{3}_Flow{2}")=HiField(16,2)	
   	SmartTags("DB_MouldEditor_HMI_uData_arShotSet{3}_Flow{3}")=HiField(16,3)
   	SmartTags("DB_MouldEditor_HMI_uData_arShotSet{3}_Flow{4}")=HiField(16,4)
   	SmartTags("DB_MouldEditor_HMI_uData_arShotSet{3}_Flow{5}")=HiField(16,5)	
   	SmartTags("DB_MouldEditor_HMI_uData_arShotSet{3}_Flow{6}")=HiField(16,6)
   	
   	SmartTags("DB_MouldEditor_HMI_uData_arShotSet{4}_Flow{1}")=HiField(21,1)
   	SmartTags("DB_MouldEditor_HMI_uData_arShotSet{4}_Flow{2}")=HiField(21,2)	
   	SmartTags("DB_MouldEditor_HMI_uData_arShotSet{4}_Flow{3}")=HiField(21,3)
   	SmartTags("DB_MouldEditor_HMI_uData_arShotSet{4}_Flow{4}")=HiField(21,4)
   	SmartTags("DB_MouldEditor_HMI_uData_arShotSet{4}_Flow{5}")=HiField(21,5)	
   	SmartTags("DB_MouldEditor_HMI_uData_arShotSet{4}_Flow{6}")=HiField(21,6)
   	
   	SmartTags("DB_MouldEditor_HMI_uData_arShotSet{5}_Flow{1}")=HiField(26,1)
   	SmartTags("DB_MouldEditor_HMI_uData_arShotSet{5}_Flow{2}")=HiField(26,2)	
   	SmartTags("DB_MouldEditor_HMI_uData_arShotSet{5}_Flow{3}")=HiField(26,3)
   	SmartTags("DB_MouldEditor_HMI_uData_arShotSet{5}_Flow{4}")=HiField(26,4)
   	SmartTags("DB_MouldEditor_HMI_uData_arShotSet{5}_Flow{5}")=HiField(26,5)	
   	SmartTags("DB_MouldEditor_HMI_uData_arShotSet{5}_Flow{6}")=HiField(26,6)
   	
   	SmartTags("DB_MouldEditor_HMI_uData_arShotSet{6}_Flow{1}")=HiField(31,1)
   	SmartTags("DB_MouldEditor_HMI_uData_arShotSet{6}_Flow{2}")=HiField(31,2)	
   	SmartTags("DB_MouldEditor_HMI_uData_arShotSet{6}_Flow{3}")=HiField(31,3)
   	SmartTags("DB_MouldEditor_HMI_uData_arShotSet{6}_Flow{4}")=HiField(31,4)
   	SmartTags("DB_MouldEditor_HMI_uData_arShotSet{6}_Flow{5}")=HiField(31,5)	
   	SmartTags("DB_MouldEditor_HMI_uData_arShotSet{6}_Flow{6}")=HiField(31,6)
   	
   	SmartTags("DB_MouldEditor_HMI_uData_arShotSet{7}_Flow{1}")=HiField(36,1)
   	SmartTags("DB_MouldEditor_HMI_uData_arShotSet{7}_Flow{2}")=HiField(36,2)	
   	SmartTags("DB_MouldEditor_HMI_uData_arShotSet{7}_Flow{3}")=HiField(36,3)
   	SmartTags("DB_MouldEditor_HMI_uData_arShotSet{7}_Flow{4}")=HiField(36,4)
   	SmartTags("DB_MouldEditor_HMI_uData_arShotSet{7}_Flow{5}")=HiField(36,5)	
   	SmartTags("DB_MouldEditor_HMI_uData_arShotSet{7}_Flow{6}")=HiField(36,6)
   	
   	SmartTags("DB_MouldEditor_HMI_uData_arShotSet{8}_Flow{1}")=HiField(41,1)
   	SmartTags("DB_MouldEditor_HMI_uData_arShotSet{8}_Flow{2}")=HiField(41,2)	
   	SmartTags("DB_MouldEditor_HMI_uData_arShotSet{8}_Flow{3}")=HiField(41,3)
   	SmartTags("DB_MouldEditor_HMI_uData_arShotSet{8}_Flow{4}")=HiField(41,4)
   	SmartTags("DB_MouldEditor_HMI_uData_arShotSet{8}_Flow{5}")=HiField(41,5)	
   	SmartTags("DB_MouldEditor_HMI_uData_arShotSet{8}_Flow{6}")=HiField(41,6)
   	
   	'//PRESSURE
   	SmartTags("DB_MouldEditor_HMI_uData_arShotSet{1}_Pressure{1}")=HiField(7,1)
   	SmartTags("DB_MouldEditor_HMI_uData_arShotSet{1}_Pressure{2}")=HiField(7,2)
   	SmartTags("DB_MouldEditor_HMI_uData_arShotSet{1}_Pressure{3}")=HiField(7,3)
   	SmartTags("DB_MouldEditor_HMI_uData_arShotSet{1}_Pressure{4}")=HiField(7,4)
   	SmartTags("DB_MouldEditor_HMI_uData_arShotSet{1}_Pressure{5}")=HiField(7,5)
   	SmartTags("DB_MouldEditor_HMI_uData_arShotSet{1}_Pressure{6}")=HiField(7,6)
   	
   	SmartTags("DB_MouldEditor_HMI_uData_arShotSet{2}_Pressure{1}")=HiField(12,1)
   	SmartTags("DB_MouldEditor_HMI_uData_arShotSet{2}_Pressure{2}")=HiField(12,2)
   	SmartTags("DB_MouldEditor_HMI_uData_arShotSet{2}_Pressure{3}")=HiField(12,3)
   	SmartTags("DB_MouldEditor_HMI_uData_arShotSet{2}_Pressure{4}")=HiField(12,4)
   	SmartTags("DB_MouldEditor_HMI_uData_arShotSet{2}_Pressure{5}")=HiField(12,5)
   	SmartTags("DB_MouldEditor_HMI_uData_arShotSet{2}_Pressure{6}")=HiField(12,6)
   	
   	SmartTags("DB_MouldEditor_HMI_uData_arShotSet{3}_Pressure{1}")=HiField(17,1)
   	SmartTags("DB_MouldEditor_HMI_uData_arShotSet{3}_Pressure{2}")=HiField(17,2)
   	SmartTags("DB_MouldEditor_HMI_uData_arShotSet{3}_Pressure{3}")=HiField(17,3)
   	SmartTags("DB_MouldEditor_HMI_uData_arShotSet{3}_Pressure{4}")=HiField(17,4)
   	SmartTags("DB_MouldEditor_HMI_uData_arShotSet{3}_Pressure{5}")=HiField(17,5)
   	SmartTags("DB_MouldEditor_HMI_uData_arShotSet{3}_Pressure{6}")=HiField(17,6)
   	
   	SmartTags("DB_MouldEditor_HMI_uData_arShotSet{4}_Pressure{1}")=HiField(22,1)
   	SmartTags("DB_MouldEditor_HMI_uData_arShotSet{4}_Pressure{2}")=HiField(22,2)
   	SmartTags("DB_MouldEditor_HMI_uData_arShotSet{4}_Pressure{3}")=HiField(22,3)
   	SmartTags("DB_MouldEditor_HMI_uData_arShotSet{4}_Pressure{4}")=HiField(22,4)
   	SmartTags("DB_MouldEditor_HMI_uData_arShotSet{4}_Pressure{5}")=HiField(22,5)
   	SmartTags("DB_MouldEditor_HMI_uData_arShotSet{4}_Pressure{6}")=HiField(22,6)
   	
   	SmartTags("DB_MouldEditor_HMI_uData_arShotSet{5}_Pressure{1}")=HiField(27,1)
   	SmartTags("DB_MouldEditor_HMI_uData_arShotSet{5}_Pressure{2}")=HiField(27,2)
   	SmartTags("DB_MouldEditor_HMI_uData_arShotSet{5}_Pressure{3}")=HiField(27,3)
   	SmartTags("DB_MouldEditor_HMI_uData_arShotSet{5}_Pressure{4}")=HiField(27,4)
   	SmartTags("DB_MouldEditor_HMI_uData_arShotSet{5}_Pressure{5}")=HiField(27,5)
   	SmartTags("DB_MouldEditor_HMI_uData_arShotSet{5}_Pressure{6}")=HiField(27,6)
   	
   	SmartTags("DB_MouldEditor_HMI_uData_arShotSet{6}_Pressure{1}")=HiField(32,1)
   	SmartTags("DB_MouldEditor_HMI_uData_arShotSet{6}_Pressure{2}")=HiField(32,2)
   	SmartTags("DB_MouldEditor_HMI_uData_arShotSet{6}_Pressure{3}")=HiField(32,3)
   	SmartTags("DB_MouldEditor_HMI_uData_arShotSet{6}_Pressure{4}")=HiField(32,4)
   	SmartTags("DB_MouldEditor_HMI_uData_arShotSet{6}_Pressure{5}")=HiField(32,5)
   	SmartTags("DB_MouldEditor_HMI_uData_arShotSet{6}_Pressure{6}")=HiField(32,6)
   	
